REGION Network 18
   RUNG wire#powerrail
      Contact( "PanelCompBAJA MTA".MantMC062 )
      { S7_GenerateENO := "TRUE" } Move(in := 0, out1 => "CmpBajaAuto".MenuMC062)
      wire#w1
      Coil( "Tag_6" )
   END_RUNG
   RUNG wire#powerrail
      I_Contact( "PanelCompBAJA MTA".MantMC062 )
      Contact( "CmpBajaAuto".AutoMC062 )
      { S7_GenerateENO := "TRUE" } Move(in := 1, out1 => "CmpBajaAuto".MenuMC062)
   END_RUNG wire#w1
   RUNG wire#powerrail
      I_Contact( "PanelCompBAJA MTA".MantMC062 )
      I_Contact( "CmpBajaAuto".AutoMC062 )
      { S7_GenerateENO := "TRUE" } Move(in := 2, out1 => "CmpBajaAuto".MenuMC062)
   END_RUNG wire#w1
   // the same network as SCL:
   // ENO of a box is taken as its EN; it also drops when the box reports an error
   IF "PanelCompBAJA MTA".MantMC062 THEN "CmpBajaAuto".MenuMC062 := 0; END_IF;
   #_w1 := NOT "PanelCompBAJA MTA".MantMC062 AND "CmpBajaAuto".AutoMC062;
   IF #_w1 THEN "CmpBajaAuto".MenuMC062 := 1; END_IF;
   #_w2 := NOT "PanelCompBAJA MTA".MantMC062 AND NOT "CmpBajaAuto".AutoMC062;
   IF #_w2 THEN "CmpBajaAuto".MenuMC062 := 2; END_IF;
   "Tag_6" := "PanelCompBAJA MTA".MantMC062 OR #_w1 OR #_w2;
END_REGION

REGION Network 19
   RUNG wire#powerrail
      Contact( "PanelCompBAJA MTA".MantMC063 )
      { S7_GenerateENO := "TRUE" } Move(in := 0, out1 => "CmpBajaAuto".MenuMC063)
      wire#w1
      Coil( "Tag_6" )
   END_RUNG
   RUNG wire#powerrail
      I_Contact( "PanelCompBAJA MTA".MantMC063 )
      Contact( "CmpBajaAuto".AutoMC063 )
      { S7_GenerateENO := "TRUE" } Move(in := 1, out1 => "CmpBajaAuto".MenuMC063)
   END_RUNG wire#w1
   RUNG wire#powerrail
      I_Contact( "PanelCompBAJA MTA".MantMC063 )
      I_Contact( "CmpBajaAuto".AutoMC063 )
      { S7_GenerateENO := "TRUE" } Move(in := 2, out1 => "CmpBajaAuto".MenuMC063)
   END_RUNG wire#w1
   // the same network as SCL:
   // ENO of a box is taken as its EN; it also drops when the box reports an error
   IF "PanelCompBAJA MTA".MantMC063 THEN "CmpBajaAuto".MenuMC063 := 0; END_IF;
   #_w1 := NOT "PanelCompBAJA MTA".MantMC063 AND "CmpBajaAuto".AutoMC063;
   IF #_w1 THEN "CmpBajaAuto".MenuMC063 := 1; END_IF;
   #_w2 := NOT "PanelCompBAJA MTA".MantMC063 AND NOT "CmpBajaAuto".AutoMC063;
   IF #_w2 THEN "CmpBajaAuto".MenuMC063 := 2; END_IF;
   "Tag_6" := "PanelCompBAJA MTA".MantMC063 OR #_w1 OR #_w2;
END_REGION

REGION Network 20
   RUNG wire#powerrail
      Contact( "PanelCompBAJA MTA".MantMC064 )
      { S7_GenerateENO := "TRUE" } Move(in := 0, out1 => "CmpBajaAuto".MenuMC064)
      wire#w1
      Coil( "Tag_6" )
   END_RUNG
   RUNG wire#powerrail
      I_Contact( "PanelCompBAJA MTA".MantMC064 )
      Contact( "CmpBajaAuto".AutoMC064 )
      { S7_GenerateENO := "TRUE" } Move(in := 1, out1 => "CmpBajaAuto".MenuMC064)
   END_RUNG wire#w1
   RUNG wire#powerrail
      I_Contact( "PanelCompBAJA MTA".MantMC064 )
      I_Contact( "CmpBajaAuto".AutoMC064 )
      { S7_GenerateENO := "TRUE" } Move(in := 2, out1 => "CmpBajaAuto".MenuMC064)
   END_RUNG wire#w1
   // the same network as SCL:
   // ENO of a box is taken as its EN; it also drops when the box reports an error
   IF "PanelCompBAJA MTA".MantMC064 THEN "CmpBajaAuto".MenuMC064 := 0; END_IF;
   #_w1 := NOT "PanelCompBAJA MTA".MantMC064 AND "CmpBajaAuto".AutoMC064;
   IF #_w1 THEN "CmpBajaAuto".MenuMC064 := 1; END_IF;
   #_w2 := NOT "PanelCompBAJA MTA".MantMC064 AND NOT "CmpBajaAuto".AutoMC064;
   IF #_w2 THEN "CmpBajaAuto".MenuMC064 := 2; END_IF;
   "Tag_6" := "PanelCompBAJA MTA".MantMC064 OR #_w1 OR #_w2;
END_REGION
END_FUNCTION

// folder: Entradas Analógicas

FUNCTION "LecturasAnalógicasMTA" : Void   // FC15, LAD
{ S7_Optimized_Access := 'FALSE' }
VERSION : 0.1
BEGIN

REGION Network 1: Lectura Temperatura Torres Cavaleto
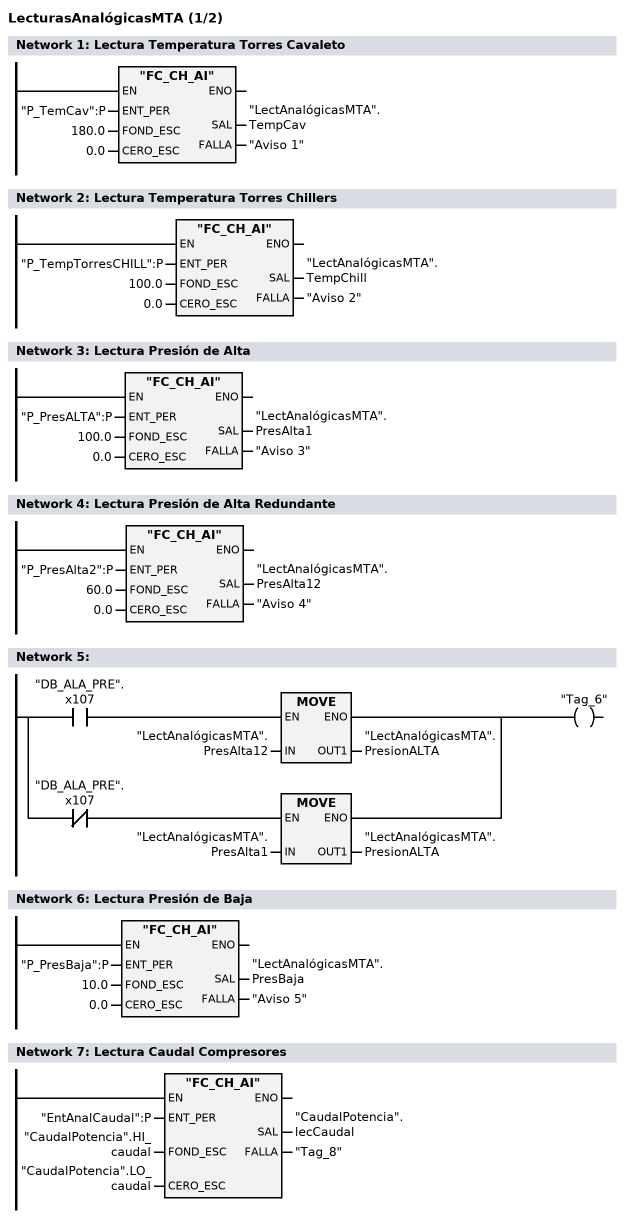
   RUNG wire#powerrail
      "FC_CH_AI"(ENT_PER := "P_TemCav":P, FOND_ESC := 180.0, CERO_ESC := 0.0, SAL => "LectAnalógicasMTA".TempCav, FALLA => "Aviso 1")
   END_RUNG
   // the same network as SCL:
   "FC_CH_AI"(ENT_PER := "P_TemCav":P,
              FOND_ESC := 180.0,
              CERO_ESC := 0.0,
              SAL => "LectAnalógicasMTA".TempCav,
              FALLA => "Aviso 1");
END_REGION

REGION Network 2: Lectura Temperatura Torres Chillers
   RUNG wire#powerrail
      "FC_CH_AI"(ENT_PER := "P_TempTorresCHILL":P, FOND_ESC := 100.0, CERO_ESC := 0.0, SAL => "LectAnalógicasMTA".TempChill, FALLA => "Aviso 2")
   END_RUNG
   // the same network as SCL:
   "FC_CH_AI"(ENT_PER := "P_TempTorresCHILL":P,
              FOND_ESC := 100.0,
              CERO_ESC := 0.0,
              SAL => "LectAnalógicasMTA".TempChill,
              FALLA => "Aviso 2");
END_REGION

REGION Network 3: Lectura Presión de Alta
   RUNG wire#powerrail
      "FC_CH_AI"(ENT_PER := "P_PresALTA":P, FOND_ESC := 100.0, CERO_ESC := 0.0, SAL => "LectAnalógicasMTA".PresAlta1, FALLA => "Aviso 3")
   END_RUNG
   // the same network as SCL:
   "FC_CH_AI"(ENT_PER := "P_PresALTA":P,
              FOND_ESC := 100.0,
              CERO_ESC := 0.0,
              SAL => "LectAnalógicasMTA".PresAlta1,
              FALLA => "Aviso 3");
END_REGION

REGION Network 4: Lectura Presión de Alta Redundante
   RUNG wire#powerrail
      "FC_CH_AI"(ENT_PER := "P_PresAlta2":P, FOND_ESC := 60.0, CERO_ESC := 0.0, SAL => "LectAnalógicasMTA".PresAlta12, FALLA => "Aviso 4")
   END_RUNG
   // the same network as SCL:
   "FC_CH_AI"(ENT_PER := "P_PresAlta2":P,
              FOND_ESC := 60.0,
              CERO_ESC := 0.0,
              SAL => "LectAnalógicasMTA".PresAlta12,
              FALLA => "Aviso 4");
END_REGION

REGION Network 5
   RUNG wire#powerrail
      Contact( "DB_ALA_PRE".x107 )
      { S7_GenerateENO := "TRUE" } Move(in := "LectAnalógicasMTA".PresAlta12, out1 => "LectAnalógicasMTA".PresionALTA)
      wire#w1
      Coil( "Tag_6" )
   END_RUNG
   RUNG wire#powerrail
      I_Contact( "DB_ALA_PRE".x107 )
      { S7_GenerateENO := "TRUE" } Move(in := "LectAnalógicasMTA".PresAlta1, out1 => "LectAnalógicasMTA".PresionALTA)
   END_RUNG wire#w1
   // the same network as SCL:
   // ENO of a box is taken as its EN; it also drops when the box reports an error
   IF "DB_ALA_PRE".x107 THEN "LectAnalógicasMTA".PresionALTA := "LectAnalógicasMTA".PresAlta12; END_IF;
   IF NOT "DB_ALA_PRE".x107 THEN "LectAnalógicasMTA".PresionALTA := "LectAnalógicasMTA".PresAlta1; END_IF;
   "Tag_6" := "DB_ALA_PRE".x107 OR NOT "DB_ALA_PRE".x107;
END_REGION

REGION Network 6: Lectura Presión de Baja
   RUNG wire#powerrail
      "FC_CH_AI"(ENT_PER := "P_PresBaja":P, FOND_ESC := 10.0, CERO_ESC := 0.0, SAL => "LectAnalógicasMTA".PresBaja, FALLA => "Aviso 5")
   END_RUNG
   // the same network as SCL:
   "FC_CH_AI"(ENT_PER := "P_PresBaja":P,
              FOND_ESC := 10.0,
              CERO_ESC := 0.0,
              SAL => "LectAnalógicasMTA".PresBaja,
              FALLA => "Aviso 5");
END_REGION

REGION Network 7: Lectura Caudal Compresores
   RUNG wire#powerrail
      "FC_CH_AI"(ENT_PER := "EntAnalCaudal":P, FOND_ESC := "CaudalPotencia".HI_caudal, CERO_ESC := "CaudalPotencia".LO_caudal, SAL => "CaudalPotencia".lecCaudal, FALLA => "Tag_8")
   END_RUNG
   // the same network as SCL:
   "FC_CH_AI"(ENT_PER := "EntAnalCaudal":P,
              FOND_ESC := "CaudalPotencia".HI_caudal,
              CERO_ESC := "CaudalPotencia".LO_caudal,
              SAL => "CaudalPotencia".lecCaudal,
              FALLA => "Tag_8");
END_REGION

REGION Network 8: Lectura Potencia Compresores
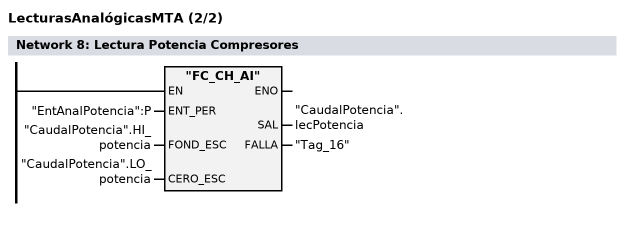
   RUNG wire#powerrail
      "FC_CH_AI"(ENT_PER := "EntAnalPotencia":P, FOND_ESC := "CaudalPotencia".HI_potencia, CERO_ESC := "CaudalPotencia".LO_potencia, SAL => "CaudalPotencia".lecPotencia, FALLA => "Tag_16")
   END_RUNG
   // the same network as SCL:
   "FC_CH_AI"(ENT_PER := "EntAnalPotencia":P,
              FOND_ESC := "CaudalPotencia".HI_potencia,
              CERO_ESC := "CaudalPotencia".LO_potencia,
              SAL => "CaudalPotencia".lecPotencia,
              FALLA => "Tag_16");
END_REGION
END_FUNCTION

// folder: Horas de Marcha

ORGANIZATION_BLOCK "CYC_INT5"   // OB35, LAD
{ S7_Optimized_Access := 'FALSE' }
VERSION : 0.1
   VAR_TEMP   // added for the SCL form of the ladder/FBD networks
      _w1 : Bool;
      _w2 : Bool;
      _w3 : Bool;
      _w4 : Bool;
   END_VAR
BEGIN

REGION Network 1 (STL)
         A     "MC001";
         A     "MC001-CO";
         =     <??.?>;
         A     <??.?>;
         A(;
         L     "SumaOB35 MTA".SMMC001;
         L     600;
         <I;
         );
         JNB   M001;
         L     1;
         L     "SumaOB35 MTA".SMMC001;
         +D;
         T     "SumaOB35 MTA".SMMC001;
   M001: NOP   0;
         A     <??.?>;
         A(;
         L     "SumaOB35 MTA".SMMC001;
         L     600;
         >=I;
         );
         =     <??.?>;
         A     <??.?>;
         JNB   M002;
         L     1;
         L     "SumaOB35 MTA".MMMC001;
         +D;
         T     "SumaOB35 MTA".MMMC001;
   M002: NOP   0;
         A     <??.?>;
         JNB   M003;
         L     0;
         T     "SumaOB35 MTA".SMMC001;
   M003: NOP   0;
         A     <??.?>;
         A(;
         L     "SumaOB35 MTA".MMMC001;
         L     60;
         >=I;
         );
         =     <??.?>;
         A     <??.?>;
         JNB   M004;
         L     1;
         L     "SumaOB35 MTA".HMMC001;
         +D;
         T     "SumaOB35 MTA".HMMC001;
   M004: NOP   0;
         A     <??.?>;
         JNB   M005;
         L     0;
         T     "SumaOB35 MTA".MMMC001;
   M005: NOP   0;
END_REGION

REGION Network 2 (STL)
         A     "MC002";
         A     "MC002-CO";
         =     <??.?>;
         A     <??.?>;
         A(;
         L     "SumaOB35 MTA".SMMC002;
         L     600;
         <I;
         );
         JNB   M006;
         L     1;
         L     "SumaOB35 MTA".SMMC002;
         +D;
         T     "SumaOB35 MTA".SMMC002;
   M006: NOP   0;
         A     <??.?>;
         A(;
         L     "SumaOB35 MTA".SMMC002;
         L     600;
         >=I;
         );
         =     <??.?>;
         A     <??.?>;
         JNB   M007;
         L     1;
         L     "SumaOB35 MTA".MMMC002;
         +D;
         T     "SumaOB35 MTA".MMMC002;
   M007: NOP   0;
         A     <??.?>;
         JNB   M008;
         L     0;
         T     "SumaOB35 MTA".SMMC002;
   M008: NOP   0;
         A     <??.?>;
         A(;
         L     "SumaOB35 MTA".MMMC002;
         L     60;
         >=I;
         );
         =     <??.?>;
         A     <??.?>;
         JNB   M009;
         L     1;
         L     "SumaOB35 MTA".HMMC002;
         +D;
         T     "SumaOB35 MTA".HMMC002;
   M009: NOP   0;
         A     <??.?>;
         JNB   M00a;
         L     0;
         T     "SumaOB35 MTA".MMMC002;
   M00a: NOP   0;
END_REGION

REGION Network 3 (STL)
         A     "MC003";
         A     "MC003-CO";
         =     <??.?>;
         A     <??.?>;
         A(;
         L     "SumaOB35 MTA".SMMC003;
         L     600;
         <I;
         );
         JNB   M00b;
         L     1;
         L     "SumaOB35 MTA".SMMC003;
         +D;
         T     "SumaOB35 MTA".SMMC003;
   M00b: NOP   0;
         A     <??.?>;
         A(;
         L     "SumaOB35 MTA".SMMC003;
         L     600;
         >=I;
         );
         =     <??.?>;
         A     <??.?>;
         JNB   M00c;
         L     1;
         L     "SumaOB35 MTA".MMMC003;
         +D;
         T     "SumaOB35 MTA".MMMC003;
   M00c: NOP   0;
         A     <??.?>;
         JNB   M00d;
         L     0;
         T     "SumaOB35 MTA".SMMC003;
   M00d: NOP   0;
         A     <??.?>;
         A(;
         L     "SumaOB35 MTA".MMMC003;
         L     60;
         >=I;
         );
         =     <??.?>;
         A     <??.?>;
         JNB   M00e;
         L     1;
         L     "SumaOB35 MTA".HMMC003;
         +D;
         T     "SumaOB35 MTA".HMMC003;
   M00e: NOP   0;
         A     <??.?>;
         JNB   M00f;
         L     0;
         T     "SumaOB35 MTA".MMMC003;
   M00f: NOP   0;
END_REGION

REGION Network 4 (STL)
         A     "MC004";
         A     "MC004-CO";
         =     <??.?>;
         A     <??.?>;
         A(;
         L     "SumaOB35 MTA".SMMC004;
         L     600;
         <I;
         );
         JNB   M010;
         L     1;
         L     "SumaOB35 MTA".SMMC004;
         +D;
         T     "SumaOB35 MTA".SMMC004;
   M010: NOP   0;
         A     <??.?>;
         A(;
         L     "SumaOB35 MTA".SMMC004;
         L     600;
         >=I;
         );
         =     <??.?>;
         A     <??.?>;
         JNB   M011;
         L     1;
         L     "SumaOB35 MTA".MMMC004;
         +D;
         T     "SumaOB35 MTA".MMMC004;
   M011: NOP   0;
         A     <??.?>;
         JNB   M012;
         L     0;
         T     "SumaOB35 MTA".SMMC004;
   M012: NOP   0;
         A     <??.?>;
         A(;
         L     "SumaOB35 MTA".MMMC004;
         L     60;
         >=I;
         );
         =     <??.?>;
         A     <??.?>;
         JNB   M013;
         L     1;
         L     "SumaOB35 MTA".HMMC004;
         +D;
         T     "SumaOB35 MTA".HMMC004;
   M013: NOP   0;
         A     <??.?>;
         JNB   M014;
         L     0;
         T     "SumaOB35 MTA".MMMC004;
   M014: NOP   0;
END_REGION

REGION Network 5 (STL)
         A     "MC005";
         A     "MC005-CO";
         =     <??.?>;
         A     <??.?>;
         A(;
         L     "SumaOB35 MTA".SMMC005;
         L     600;
         <I;
         );
         JNB   M015;
         L     1;
         L     "SumaOB35 MTA".SMMC005;
         +D;
         T     "SumaOB35 MTA".SMMC005;
   M015: NOP   0;
         A     <??.?>;
         A(;
         L     "SumaOB35 MTA".SMMC005;
         L     600;
         >=I;
         );
         =     <??.?>;
         A     <??.?>;
         JNB   M016;
         L     1;
         L     "SumaOB35 MTA".MMMC005;
         +D;
         T     "SumaOB35 MTA".MMMC005;
   M016: NOP   0;
         A     <??.?>;
         JNB   M017;
         L     0;
         T     "SumaOB35 MTA".SMMC005;
   M017: NOP   0;
         A     <??.?>;
         A(;
         L     "SumaOB35 MTA".MMMC005;
         L     60;
         >=I;
         );
         =     <??.?>;
         A     <??.?>;
         JNB   M018;
         L     1;
         L     "SumaOB35 MTA".HMMC005;
         +D;
         T     "SumaOB35 MTA".HMMC005;
   M018: NOP   0;
         A     <??.?>;
         JNB   M019;
         L     0;
         T     "SumaOB35 MTA".MMMC005;
   M019: NOP   0;
END_REGION

REGION Network 6 (STL)
         A     "MC006";
         A     "MC006-CO";
         =     <??.?>;
         A     <??.?>;
         A(;
         L     "SumaOB35 MTA".SMMC006;
         L     600;
         <I;
         );
         JNB   M020;
         L     1;
         L     "SumaOB35 MTA".SMMC006;
         +D;
         T     "SumaOB35 MTA".SMMC006;
   M020: NOP   0;
         A     <??.?>;
         A(;
         L     "SumaOB35 MTA".SMMC006;
         L     600;
         >=I;
         );
         =     <??.?>;
         A     <??.?>;
         JNB   M021;
         L     1;
         L     "SumaOB35 MTA".MMMC006;
         +D;
         T     "SumaOB35 MTA".MMMC006;
   M021: NOP   0;
         A     <??.?>;
         JNB   M022;
         L     0;
         T     "SumaOB35 MTA".SMMC006;
   M022: NOP   0;
         A     <??.?>;
         A(;
         L     "SumaOB35 MTA".MMMC006;
         L     60;
         >=I;
         );
         =     <??.?>;
         A     <??.?>;
         JNB   M023;
         L     1;
         L     "SumaOB35 MTA".HMMC006;
         +D;
         T     "SumaOB35 MTA".HMMC006;
   M023: NOP   0;
         A     <??.?>;
         JNB   M024;
         L     0;
         T     "SumaOB35 MTA".MMMC006;
   M024: NOP   0;
END_REGION

REGION Network 7: Encendido de PLC
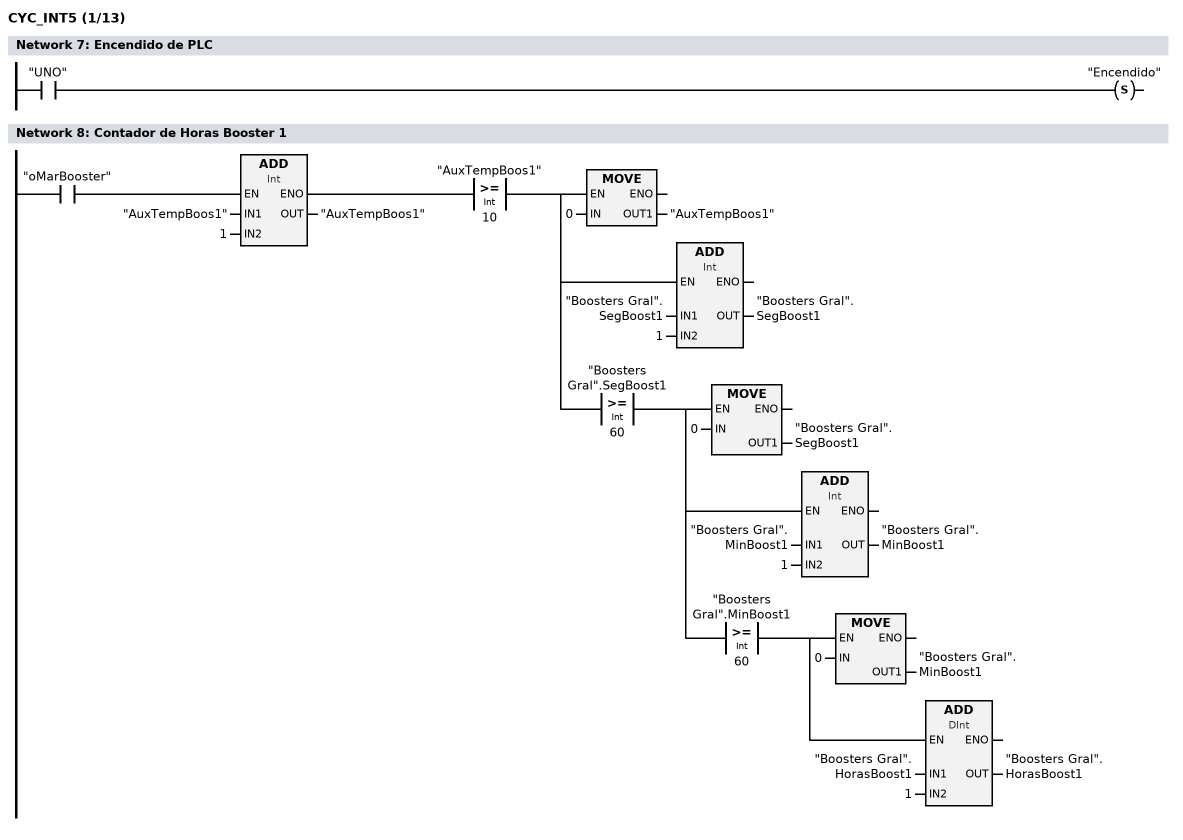
   RUNG wire#powerrail
      Contact( "UNO" )
      S_Coil( "Encendido" )
   END_RUNG
   // the same network as SCL:
   IF "UNO" THEN "Encendido" := TRUE; END_IF;
END_REGION

REGION Network 8: Contador de Horas Booster 1
   RUNG wire#powerrail
      Contact( "oMarBooster" )
      { S7_Templates := "SrcType := Int"; S7_GenerateENO := "TRUE" } Add(in1 := "AuxTempBoos1", in2 := 1, out => "AuxTempBoos1")
      { S7_Templates := "SrcType := Int" } GE_Contact(in1 := "AuxTempBoos1", in2 := 10)
      wire#w1
      { S7_GenerateENO := "TRUE" } Move(in := 0, out1 => "AuxTempBoos1")
   END_RUNG
   RUNG wire#w1
      { S7_Templates := "SrcType := Int"; S7_GenerateENO := "TRUE" } Add(in1 := "Boosters Gral".SegBoost1, in2 := 1, out => "Boosters Gral".SegBoost1)
   END_RUNG
   RUNG wire#w1
      { S7_Templates := "SrcType := Int" } GE_Contact(in1 := "Boosters Gral".SegBoost1, in2 := 60)
      wire#w2
      { S7_GenerateENO := "TRUE" } Move(in := 0, out1 => "Boosters Gral".SegBoost1)
   END_RUNG
   RUNG wire#w2
      { S7_Templates := "SrcType := Int"; S7_GenerateENO := "TRUE" } Add(in1 := "Boosters Gral".MinBoost1, in2 := 1, out => "Boosters Gral".MinBoost1)
   END_RUNG
   RUNG wire#w2
      { S7_Templates := "SrcType := Int" } GE_Contact(in1 := "Boosters Gral".MinBoost1, in2 := 60)
      wire#w3
      { S7_GenerateENO := "TRUE" } Move(in := 0, out1 => "Boosters Gral".MinBoost1)
   END_RUNG
   RUNG wire#w3
      { S7_Templates := "SrcType := DInt"; S7_GenerateENO := "TRUE" } Add(in1 := "Boosters Gral".HorasBoost1, in2 := 1, out => "Boosters Gral".HorasBoost1)
   END_RUNG
   // the same network as SCL:
   // ENO of a box is taken as its EN; it also drops when the box reports an error
   IF "oMarBooster" THEN "AuxTempBoos1" := "AuxTempBoos1" + 1; END_IF;
   #_w1 := "oMarBooster" AND ("AuxTempBoos1" >= 10);
   IF #_w1 THEN
       "AuxTempBoos1" := 0;
       "Boosters Gral".SegBoost1 := "Boosters Gral".SegBoost1 + 1;
   END_IF;
   #_w2 := #_w1 AND ("Boosters Gral".SegBoost1 >= 60);
   IF #_w2 THEN
       "Boosters Gral".SegBoost1 := 0;
       "Boosters Gral".MinBoost1 := "Boosters Gral".MinBoost1 + 1;
   END_IF;
   #_w3 := #_w2 AND ("Boosters Gral".MinBoost1 >= 60);
   IF #_w3 THEN
       "Boosters Gral".MinBoost1 := 0;
       "Boosters Gral".HorasBoost1 := "Boosters Gral".HorasBoost1 + 1;
   END_IF;
END_REGION

REGION Network 9: Contador de Horas Booster 2
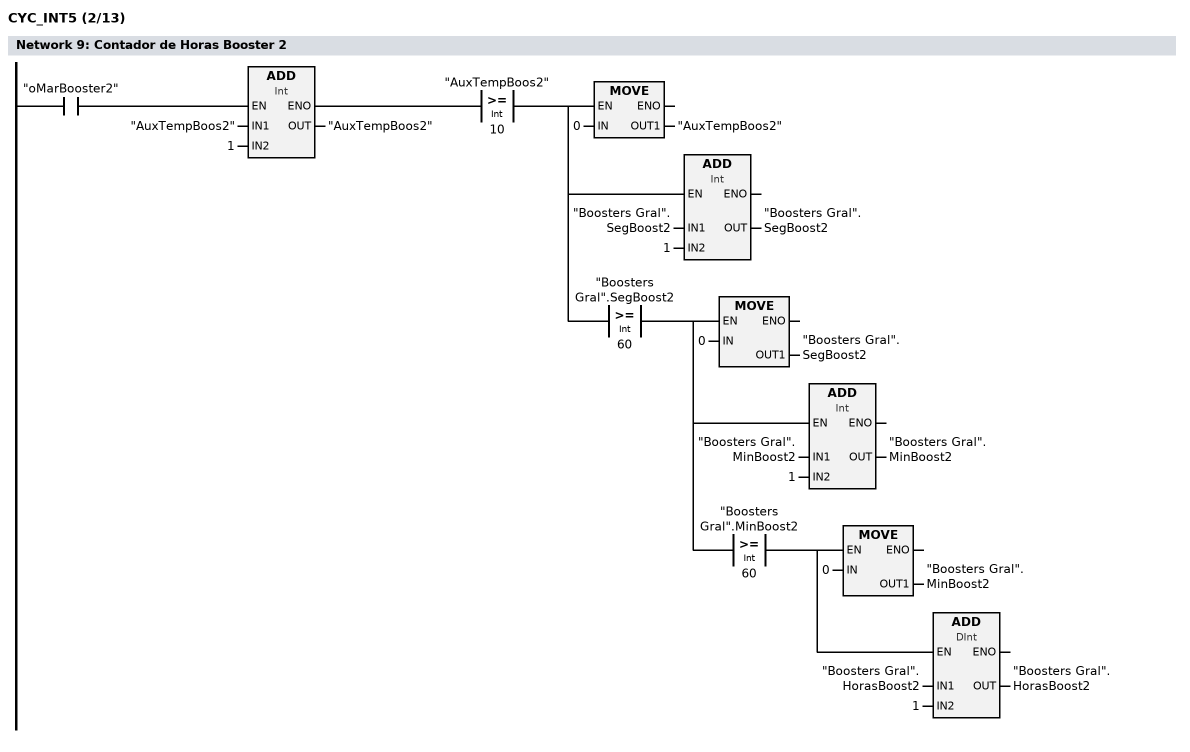
   RUNG wire#powerrail
      Contact( "oMarBooster2" )
      { S7_Templates := "SrcType := Int"; S7_GenerateENO := "TRUE" } Add(in1 := "AuxTempBoos2", in2 := 1, out => "AuxTempBoos2")
      { S7_Templates := "SrcType := Int" } GE_Contact(in1 := "AuxTempBoos2", in2 := 10)
      wire#w1
      { S7_GenerateENO := "TRUE" } Move(in := 0, out1 => "AuxTempBoos2")
   END_RUNG
   RUNG wire#w1
      { S7_Templates := "SrcType := Int"; S7_GenerateENO := "TRUE" } Add(in1 := "Boosters Gral".SegBoost2, in2 := 1, out => "Boosters Gral".SegBoost2)
   END_RUNG
   RUNG wire#w1
      { S7_Templates := "SrcType := Int" } GE_Contact(in1 := "Boosters Gral".SegBoost2, in2 := 60)
      wire#w2
      { S7_GenerateENO := "TRUE" } Move(in := 0, out1 => "Boosters Gral".SegBoost2)
   END_RUNG
   RUNG wire#w2
      { S7_Templates := "SrcType := Int"; S7_GenerateENO := "TRUE" } Add(in1 := "Boosters Gral".MinBoost2, in2 := 1, out => "Boosters Gral".MinBoost2)
   END_RUNG
   RUNG wire#w2
      { S7_Templates := "SrcType := Int" } GE_Contact(in1 := "Boosters Gral".MinBoost2, in2 := 60)
      wire#w3
      { S7_GenerateENO := "TRUE" } Move(in := 0, out1 => "Boosters Gral".MinBoost2)
   END_RUNG
   RUNG wire#w3
      { S7_Templates := "SrcType := DInt"; S7_GenerateENO := "TRUE" } Add(in1 := "Boosters Gral".HorasBoost2, in2 := 1, out => "Boosters Gral".HorasBoost2)
   END_RUNG
   // the same network as SCL:
   // ENO of a box is taken as its EN; it also drops when the box reports an error
   IF "oMarBooster2" THEN "AuxTempBoos2" := "AuxTempBoos2" + 1; END_IF;
   #_w1 := "oMarBooster2" AND ("AuxTempBoos2" >= 10);
   IF #_w1 THEN
       "AuxTempBoos2" := 0;
       "Boosters Gral".SegBoost2 := "Boosters Gral".SegBoost2 + 1;
   END_IF;
   #_w2 := #_w1 AND ("Boosters Gral".SegBoost2 >= 60);
   IF #_w2 THEN
       "Boosters Gral".SegBoost2 := 0;
       "Boosters Gral".MinBoost2 := "Boosters Gral".MinBoost2 + 1;
   END_IF;
   #_w3 := #_w2 AND ("Boosters Gral".MinBoost2 >= 60);
   IF #_w3 THEN
       "Boosters Gral".MinBoost2 := 0;
       "Boosters Gral".HorasBoost2 := "Boosters Gral".HorasBoost2 + 1;
   END_IF;
END_REGION

REGION Network 10: Horas de marcha MS050 / Contador de Horas Booster 1
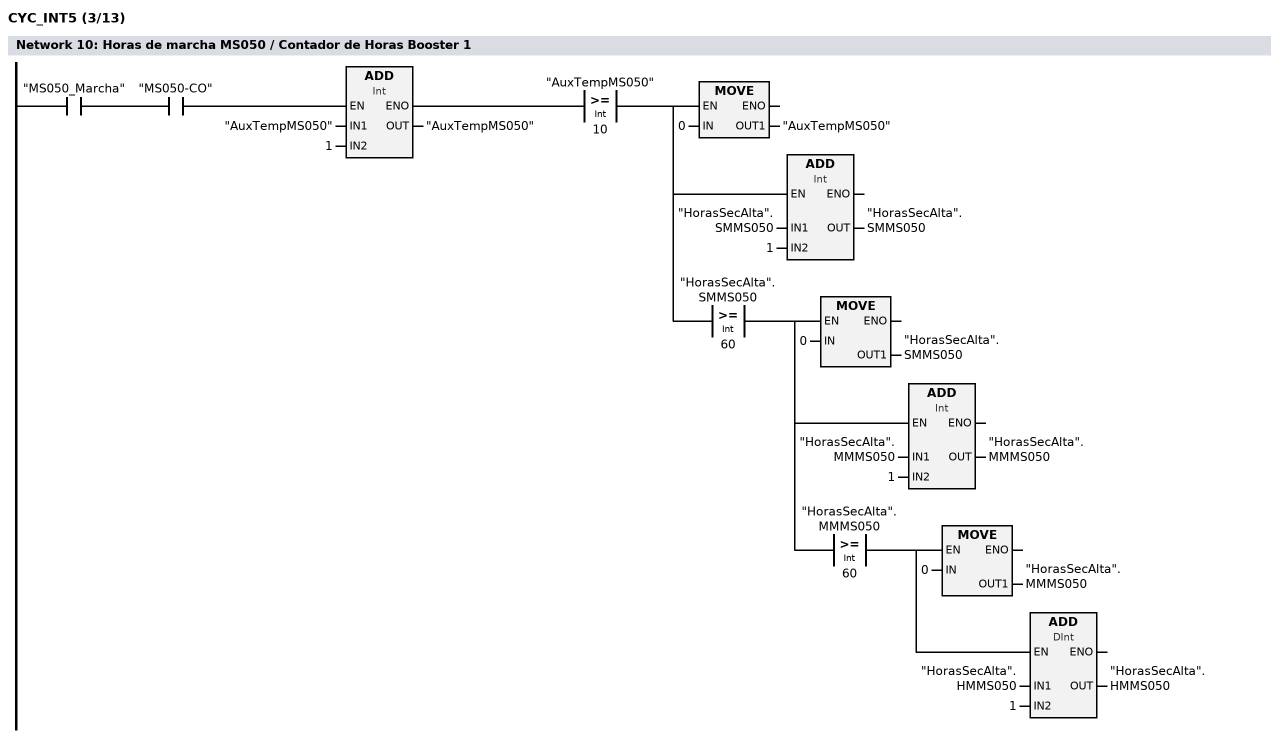
   RUNG wire#powerrail
      Contact( "MS050_Marcha" )
      Contact( "MS050-CO" )
      { S7_Templates := "SrcType := Int"; S7_GenerateENO := "TRUE" } Add(in1 := "AuxTempMS050", in2 := 1, out => "AuxTempMS050")
      { S7_Templates := "SrcType := Int" } GE_Contact(in1 := "AuxTempMS050", in2 := 10)
      wire#w1
      { S7_GenerateENO := "TRUE" } Move(in := 0, out1 => "AuxTempMS050")
   END_RUNG
   RUNG wire#w1
      { S7_Templates := "SrcType := Int"; S7_GenerateENO := "TRUE" } Add(in1 := "HorasSecAlta".SMMS050, in2 := 1, out => "HorasSecAlta".SMMS050)
   END_RUNG
   RUNG wire#w1
      { S7_Templates := "SrcType := Int" } GE_Contact(in1 := "HorasSecAlta".SMMS050, in2 := 60)
      wire#w2
      { S7_GenerateENO := "TRUE" } Move(in := 0, out1 => "HorasSecAlta".SMMS050)
   END_RUNG
   RUNG wire#w2
      { S7_Templates := "SrcType := Int"; S7_GenerateENO := "TRUE" } Add(in1 := "HorasSecAlta".MMMS050, in2 := 1, out => "HorasSecAlta".MMMS050)
   END_RUNG
   RUNG wire#w2
      { S7_Templates := "SrcType := Int" } GE_Contact(in1 := "HorasSecAlta".MMMS050, in2 := 60)
      wire#w3
      { S7_GenerateENO := "TRUE" } Move(in := 0, out1 => "HorasSecAlta".MMMS050)
   END_RUNG
   RUNG wire#w3
      { S7_Templates := "SrcType := DInt"; S7_GenerateENO := "TRUE" } Add(in1 := "HorasSecAlta".HMMS050, in2 := 1, out => "HorasSecAlta".HMMS050)
   END_RUNG
   // the same network as SCL:
   // ENO of a box is taken as its EN; it also drops when the box reports an error
   #_w1 := "MS050_Marcha" AND "MS050-CO";
   IF #_w1 THEN "AuxTempMS050" := "AuxTempMS050" + 1; END_IF;
   #_w2 := #_w1 AND ("AuxTempMS050" >= 10);
   IF #_w2 THEN
       "AuxTempMS050" := 0;
       "HorasSecAlta".SMMS050 := "HorasSecAlta".SMMS050 + 1;
   END_IF;
   #_w3 := #_w2 AND ("HorasSecAlta".SMMS050 >= 60);
   IF #_w3 THEN
       "HorasSecAlta".SMMS050 := 0;
       "HorasSecAlta".MMMS050 := "HorasSecAlta".MMMS050 + 1;
   END_IF;
   #_w4 := #_w3 AND ("HorasSecAlta".MMMS050 >= 60);
   IF #_w4 THEN
       "HorasSecAlta".MMMS050 := 0;
       "HorasSecAlta".HMMS050 := "HorasSecAlta".HMMS050 + 1;
   END_IF;
END_REGION

REGION Network 11: Horas de marcha MS051 / Contador de Horas Booster 1
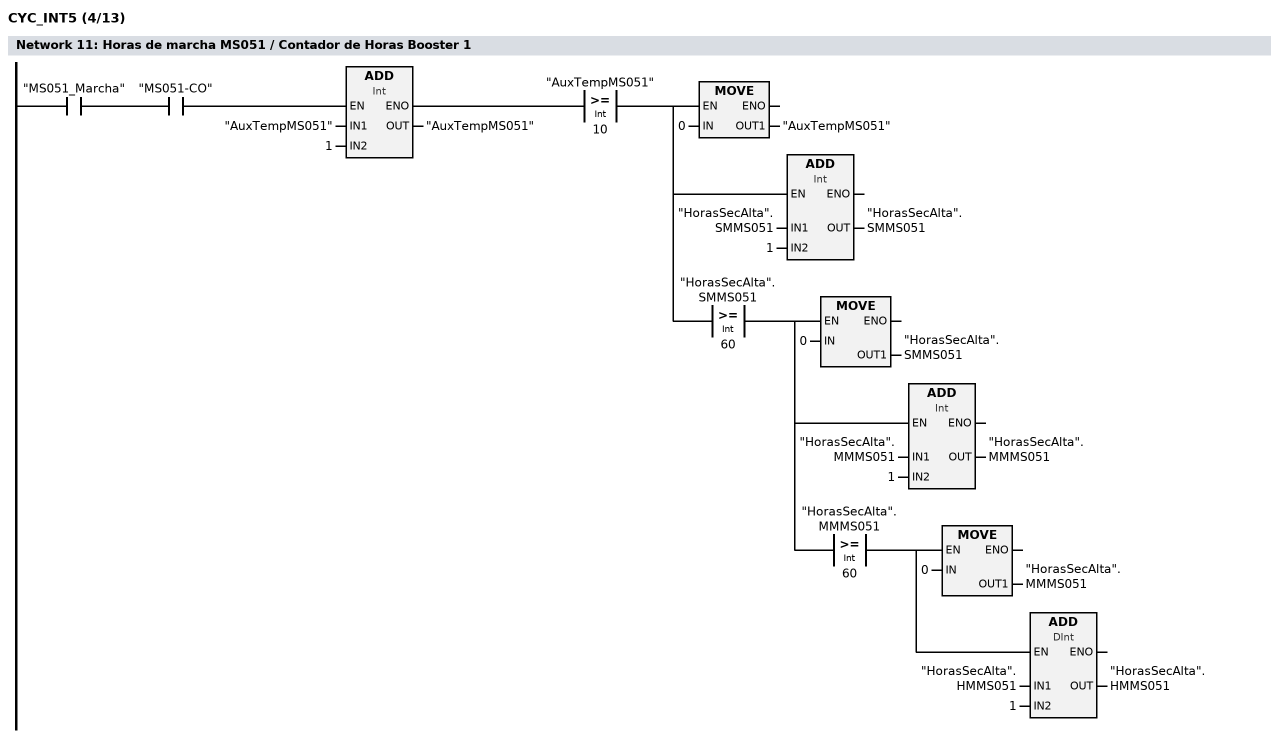
   RUNG wire#powerrail
      Contact( "MS051_Marcha" )
      Contact( "MS051-CO" )
      { S7_Templates := "SrcType := Int"; S7_GenerateENO := "TRUE" } Add(in1 := "AuxTempMS051", in2 := 1, out => "AuxTempMS051")
      { S7_Templates := "SrcType := Int" } GE_Contact(in1 := "AuxTempMS051", in2 := 10)
      wire#w1
      { S7_GenerateENO := "TRUE" } Move(in := 0, out1 => "AuxTempMS051")
   END_RUNG
   RUNG wire#w1
      { S7_Templates := "SrcType := Int"; S7_GenerateENO := "TRUE" } Add(in1 := "HorasSecAlta".SMMS051, in2 := 1, out => "HorasSecAlta".SMMS051)
   END_RUNG
   RUNG wire#w1
      { S7_Templates := "SrcType := Int" } GE_Contact(in1 := "HorasSecAlta".SMMS051, in2 := 60)
      wire#w2
      { S7_GenerateENO := "TRUE" } Move(in := 0, out1 => "HorasSecAlta".SMMS051)
   END_RUNG
   RUNG wire#w2
      { S7_Templates := "SrcType := Int"; S7_GenerateENO := "TRUE" } Add(in1 := "HorasSecAlta".MMMS051, in2 := 1, out => "HorasSecAlta".MMMS051)
   END_RUNG
   RUNG wire#w2
      { S7_Templates := "SrcType := Int" } GE_Contact(in1 := "HorasSecAlta".MMMS051, in2 := 60)
      wire#w3
      { S7_GenerateENO := "TRUE" } Move(in := 0, out1 => "HorasSecAlta".MMMS051)
   END_RUNG
   RUNG wire#w3
      { S7_Templates := "SrcType := DInt"; S7_GenerateENO := "TRUE" } Add(in1 := "HorasSecAlta".HMMS051, in2 := 1, out => "HorasSecAlta".HMMS051)
   END_RUNG
   // the same network as SCL:
   // ENO of a box is taken as its EN; it also drops when the box reports an error
   #_w1 := "MS051_Marcha" AND "MS051-CO";
   IF #_w1 THEN "AuxTempMS051" := "AuxTempMS051" + 1; END_IF;
   #_w2 := #_w1 AND ("AuxTempMS051" >= 10);
   IF #_w2 THEN
       "AuxTempMS051" := 0;
       "HorasSecAlta".SMMS051 := "HorasSecAlta".SMMS051 + 1;
   END_IF;
   #_w3 := #_w2 AND ("HorasSecAlta".SMMS051 >= 60);
   IF #_w3 THEN
       "HorasSecAlta".SMMS051 := 0;
       "HorasSecAlta".MMMS051 := "HorasSecAlta".MMMS051 + 1;
   END_IF;
   #_w4 := #_w3 AND ("HorasSecAlta".MMMS051 >= 60);
   IF #_w4 THEN
       "HorasSecAlta".MMMS051 := 0;
       "HorasSecAlta".HMMS051 := "HorasSecAlta".HMMS051 + 1;
   END_IF;
END_REGION

REGION Network 12: Horas de marcha MS052 / Contador de Horas Booster 1
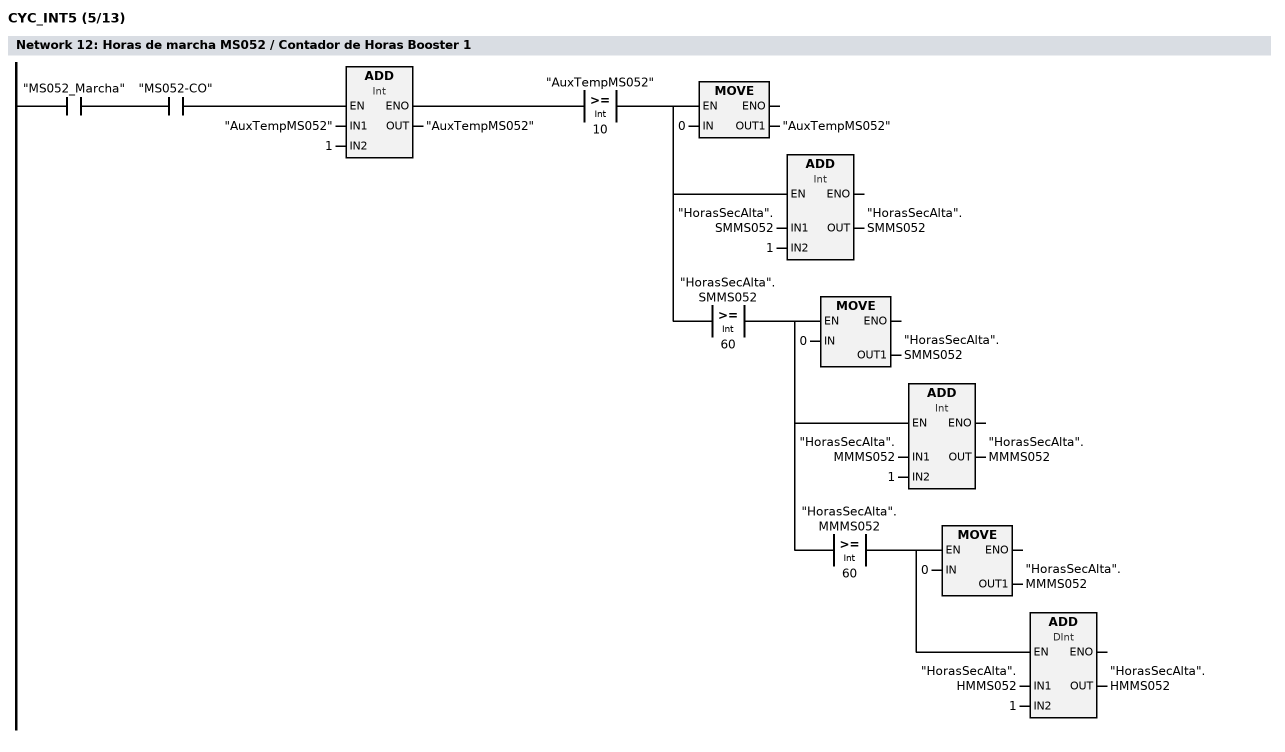
   RUNG wire#powerrail
      Contact( "MS052_Marcha" )
      Contact( "MS052-CO" )
      { S7_Templates := "SrcType := Int"; S7_GenerateENO := "TRUE" } Add(in1 := "AuxTempMS052", in2 := 1, out => "AuxTempMS052")
      { S7_Templates := "SrcType := Int" } GE_Contact(in1 := "AuxTempMS052", in2 := 10)
      wire#w1
      { S7_GenerateENO := "TRUE" } Move(in := 0, out1 => "AuxTempMS052")
   END_RUNG
   RUNG wire#w1
      { S7_Templates := "SrcType := Int"; S7_GenerateENO := "TRUE" } Add(in1 := "HorasSecAlta".SMMS052, in2 := 1, out => "HorasSecAlta".SMMS052)
   END_RUNG
   RUNG wire#w1
      { S7_Templates := "SrcType := Int" } GE_Contact(in1 := "HorasSecAlta".SMMS052, in2 := 60)
      wire#w2
      { S7_GenerateENO := "TRUE" } Move(in := 0, out1 => "HorasSecAlta".SMMS052)
   END_RUNG
   RUNG wire#w2
      { S7_Templates := "SrcType := Int"; S7_GenerateENO := "TRUE" } Add(in1 := "HorasSecAlta".MMMS052, in2 := 1, out => "HorasSecAlta".MMMS052)
   END_RUNG
   RUNG wire#w2
      { S7_Templates := "SrcType := Int" } GE_Contact(in1 := "HorasSecAlta".MMMS052, in2 := 60)
      wire#w3
      { S7_GenerateENO := "TRUE" } Move(in := 0, out1 => "HorasSecAlta".MMMS052)
   END_RUNG
   RUNG wire#w3
      { S7_Templates := "SrcType := DInt"; S7_GenerateENO := "TRUE" } Add(in1 := "HorasSecAlta".HMMS052, in2 := 1, out => "HorasSecAlta".HMMS052)
   END_RUNG
   // the same network as SCL:
   // ENO of a box is taken as its EN; it also drops when the box reports an error
   #_w1 := "MS052_Marcha" AND "MS052-CO";
   IF #_w1 THEN "AuxTempMS052" := "AuxTempMS052" + 1; END_IF;
   #_w2 := #_w1 AND ("AuxTempMS052" >= 10);
   IF #_w2 THEN
       "AuxTempMS052" := 0;
       "HorasSecAlta".SMMS052 := "HorasSecAlta".SMMS052 + 1;
   END_IF;
   #_w3 := #_w2 AND ("HorasSecAlta".SMMS052 >= 60);
   IF #_w3 THEN
       "HorasSecAlta".SMMS052 := 0;
       "HorasSecAlta".MMMS052 := "HorasSecAlta".MMMS052 + 1;
   END_IF;
   #_w4 := #_w3 AND ("HorasSecAlta".MMMS052 >= 60);
   IF #_w4 THEN
       "HorasSecAlta".MMMS052 := 0;
       "HorasSecAlta".HMMS052 := "HorasSecAlta".HMMS052 + 1;
   END_IF;
END_REGION

REGION Network 13: Horas de marcha MS053 / Contador de Horas Booster 1
